   398: 'IGG_WARNING_WORD_01_BIT_5', class IGG Warnings, trigger "62_Warning_Data_IGG_WARNING_WORD_01" bit 13
   399: 'IGG_WARNING_WORD_01_BIT_6', class IGG Warnings, trigger "62_Warning_Data_IGG_WARNING_WORD_01" bit 14
   400: 'IGG_WARNING_WORD_01_BIT_7', class IGG Warnings, trigger "62_Warning_Data_IGG_WARNING_WORD_01" bit 15
   401: 'PIT-359 INLET CSW PRESSURE - LOW', class IGG Warnings, trigger "62_Warning_Data_IGG_WARNING_WORD_02" bit 0
   402: 'PIT-359 INLET CSW PRESSURE - HIGH', class IGG Warnings, trigger "62_Warning_Data_IGG_WARNING_WORD_02" bit 1
   403: 'PIT-316 OUTLET CSW PRESSURE - LOW', class IGG Warnings, trigger "62_Warning_Data_IGG_WARNING_WORD_02" bit 2
   404: 'PIT-316 OUTLET CSW PRESSURE - HIGH', class IGG Warnings, trigger "62_Warning_Data_IGG_WARNING_WORD_02" bit 3
   405: 'PIT-316 OUTLET CSW PRESSURE - LOW LOW', class IGG Warnings, trigger "62_Warning_Data_IGG_WARNING_WORD_02" bit 4
   406: 'PIT-316 OUTLET CSW PRESSURE - HIGH HIGH', class IGG Warnings, trigger "62_Warning_Data_IGG_WARNING_WORD_02" bit 5
   407: 'IGG_WARNING_WORD_02_BIT_14', class IGG Warnings, trigger "62_Warning_Data_IGG_WARNING_WORD_02" bit 6
   408: 'IGG_WARNING_WORD_02_BIT_15', class IGG Warnings, trigger "62_Warning_Data_IGG_WARNING_WORD_02" bit 7
   409: 'PIT-102 CA PRESSURE LOW', class IGG Warnings, trigger "62_Warning_Data_IGG_WARNING_WORD_02" bit 8
   410: 'PIT-102 CA PRESSURE HIGH', class IGG Warnings, trigger "62_Warning_Data_IGG_WARNING_WORD_02" bit 9
   411: 'TIT-401 IG TEMP HIGH', class IGG Warnings, trigger "62_Warning_Data_IGG_WARNING_WORD_02" bit 10
   412: 'PIT-402 IG OUTLET PRESSURE - LOW', class IGG Warnings, trigger "62_Warning_Data_IGG_WARNING_WORD_02" bit 11
   413: 'PIT-402 IG OUTLET PRESSURE - HIGH', class IGG Warnings, trigger "62_Warning_Data_IGG_WARNING_WORD_02" bit 12
   414: 'TIT-315 SHELL CSW TEMP - HIGH', class IGG Warnings, trigger "62_Warning_Data_IGG_WARNING_WORD_02" bit 13
   415: 'TIT-319 INLET CSW TEMP - HIGH', class IGG Warnings, trigger "62_Warning_Data_IGG_WARNING_WORD_02" bit 14
   416: 'TIT-360 OUTLET CSW TEMP - HIGH', class IGG Warnings, trigger "62_Warning_Data_IGG_WARNING_WORD_02" bit 15
   417: 'FD-001 FLAME - TRIPPED', class BC Warnings, trigger "62_Warning_Data_BC_WARNING_WORD_01" bit 0
   418: 'PIT-204 FUEL OIL INLET PRESSURE - LOW LOW', class BC Warnings, trigger "62_Warning_Data_BC_WARNING_WORD_01" bit 1
   419: 'PIT-204 FUEL OIL INLET PRESSURE - LOW', class BC Warnings, trigger "62_Warning_Data_BC_WARNING_WORD_01" bit 2
   420: 'PIT-204 FUEL OIL INLET PRESSURE - HIGH', class BC Warnings, trigger "62_Warning_Data_BC_WARNING_WORD_01" bit 3
   421: 'PIT-204 FUEL OIL INLET PRESSURE - HIGH HIGH', class BC Warnings, trigger "62_Warning_Data_BC_WARNING_WORD_01" bit 4
   422: 'PIT-204 FUEL OIL INLET PRESSURE - OUT OF RANGE', class BC Warnings, trigger "62_Warning_Data_BC_WARNING_WORD_01" bit 5
   423: 'BC_WARNING_WORD_01_BIT_14', class BC Warnings, trigger "62_Warning_Data_BC_WARNING_WORD_01" bit 6
   424: 'BC_WARNING_WORD_01_BIT_15', class BC Warnings, trigger "62_Warning_Data_BC_WARNING_WORD_01" bit 7
   425: 'BC_WARNING_WORD_01_BIT_0', class BC Warnings, trigger "62_Warning_Data_BC_WARNING_WORD_01" bit 8
   426: 'PIT-204 FUEL OIL INLET PRESSURE - LOW LOW', class BC Warnings, trigger "62_Warning_Data_BC_WARNING_WORD_01" bit 9
   427: 'PIT-204 FUEL OIL INLET PRESSURE - LOW', class BC Warnings, trigger "62_Warning_Data_BC_WARNING_WORD_01" bit 10
   428: 'PIT-204 FUEL OIL INLET PRESSURE - HIGH', class BC Warnings, trigger "62_Warning_Data_BC_WARNING_WORD_01" bit 11
   429: 'PIT-204 FUEL OIL INLET PRESSURE - HIGH HIGH', class BC Warnings, trigger "62_Warning_Data_BC_WARNING_WORD_01" bit 12
   430: 'PIT-204 FUEL OIL INLET PRESSURE - OUT OF RANGE', class BC Warnings, trigger "62_Warning_Data_BC_WARNING_WORD_01" bit 13
   431: 'FD-001 FLAME NOT DETECTED', class BC Warnings, trigger "62_Warning_Data_BC_WARNING_WORD_01" bit 14
   432: 'FD-001 FLAME NOT HEALTHY', class BC Warnings, trigger "62_Warning_Data_BC_WARNING_WORD_01" bit 15
   433: 'BC_WARNING_WORD_02_BIT_8', class BC Warnings, trigger "62_Warning_Data_BC_WARNING_WORD_02" bit 0
   434: 'TIT-202 FUEL OIL INLET TEMPERATURE - LOW LOW', class BC Warnings, trigger "62_Warning_Data_BC_WARNING_WORD_02" bit 1
   435: 'TIT-202 FUEL OIL INLET TEMPERATURE - LOW', class BC Warnings, trigger "62_Warning_Data_BC_WARNING_WORD_02" bit 2
   436: 'TIT-202 FUEL OIL INLET TEMPERATURE - HIGH', class BC Warnings, trigger "62_Warning_Data_BC_WARNING_WORD_02" bit 3
   437: 'TIT-202 FUEL OIL INLET TEMPERATURE - HIGH HIGH', class BC Warnings, trigger "62_Warning_Data_BC_WARNING_WORD_02" bit 4
   438: 'TIT-202 FUEL OIL INLET TEMPERATURE - OUT OF RANGE', class BC Warnings, trigger "62_Warning_Data_BC_WARNING_WORD_02" bit 5
   439: 'BC_WARNING_WORD_02_BIT_14', class BC Warnings, trigger "62_Warning_Data_BC_WARNING_WORD_02" bit 6
   440: 'BC_WARNING_WORD_02_BIT_15', class BC Warnings, trigger "62_Warning_Data_BC_WARNING_WORD_02" bit 7
   441: 'BC_WARNING_WORD_02_BIT_0', class BC Warnings, trigger "62_Warning_Data_BC_WARNING_WORD_02" bit 8
   442: 'TIT-202 IGG INLET FUEL TEMP - LOW LOW', class BC Warnings, trigger "62_Warning_Data_BC_WARNING_WORD_02" bit 9
   443: 'TIT-202 IGG INLET FUEL TEMP - LOW', class BC Warnings, trigger "62_Warning_Data_BC_WARNING_WORD_02" bit 10
   444: 'TIT-202 IGG INLET FUEL TEMP - HIGH', class BC Warnings, trigger "62_Warning_Data_BC_WARNING_WORD_02" bit 11
   445: 'TIT-202 IGG INLET FUEL TEMP - HIGH HIGH', class BC Warnings, trigger "62_Warning_Data_BC_WARNING_WORD_02" bit 12
   446: 'TIT-202 IGG INLET FUEL TEMP - OUT OF RANGE', class BC Warnings, trigger "62_Warning_Data_BC_WARNING_WORD_02" bit 13
   447: 'BC_WARNING_WORD_02_BIT_6', class BC Warnings, trigger "62_Warning_Data_BC_WARNING_WORD_02" bit 14
   448: 'BC_WARNING_WORD_02_BIT_7', class BC Warnings, trigger "62_Warning_Data_BC_WARNING_WORD_02" bit 15
   449: 'PIT-102 CA PRESSURE - LOW LOW', class IGG Warnings, trigger "62_Warning_Data_IGG_WARNING_WORD_03" bit 0
   450: 'PIT-102 CA PRESSURE - HIGH HIGH', class IGG Warnings, trigger "62_Warning_Data_IGG_WARNING_WORD_03" bit 1
   451: 'IGG WARNING', class IGG Warnings, trigger "62_Warning_Data_IGG_WARNING_WORD_03" bit 2
   452: 'PIT-402 IG OUTLET PRESSURE - LOW LOW', class IGG Warnings, trigger "62_Warning_Data_IGG_WARNING_WORD_03" bit 3
   453: 'PIT-402 IG OUTLET PRESSURE - HIGH HIGH', class IGG Warnings, trigger "62_Warning_Data_IGG_WARNING_WORD_03" bit 4
   454: 'TIT-315 SHELL CSW TEMP - HIGH HIGH', class IGG Warnings, trigger "62_Warning_Data_IGG_WARNING_WORD_03" bit 5
   455: 'TIT-319 INLET CSW TEMP - HIGH HIGH', class IGG Warnings, trigger "62_Warning_Data_IGG_WARNING_WORD_03" bit 6
   456: 'TIT-360 OUTLET CSW TEMP - HIGH HIGH', class IGG Warnings, trigger "62_Warning_Data_IGG_WARNING_WORD_03" bit 7
   457: 'PIT-112 IA PRESSURE- OUT OF RANGE', class IGG Warnings, trigger "62_Warning_Data_IGG_WARNING_WORD_03" bit 8
   458: 'PIT-113 FUEL PRESSURE TO MAIN BURNER - OUT OF RANGE', class IGG Warnings, trigger "62_Warning_Data_IGG_WARNING_WORD_03" bit 9
   459: 'PIT-102 CA PRESSURE - OUT OF RANGE', class IGG Warnings, trigger "62_Warning_Data_IGG_WARNING_WORD_03" bit 10
   460: 'TIT-401 IG TEMP - OUT OF RANGE', class IGG Warnings, trigger "62_Warning_Data_IGG_WARNING_WORD_03" bit 11
   461: 'PIT-402 IG VENT PRESSURE - OUT OF RANGE', class IGG Warnings, trigger "62_Warning_Data_IGG_WARNING_WORD_03" bit 12
   462: 'TIT-315 SHELL CSW TEMP - OUT OF RANGE', class IGG Warnings, trigger "62_Warning_Data_IGG_WARNING_WORD_03" bit 13
   463: 'TIT-319 INLET CSW TEMP - OUT OF RANGE', class IGG Warnings, trigger "62_Warning_Data_IGG_WARNING_WORD_03" bit 14
   464: 'TIT-360 OUTLET CSW TEMP - OUT OF RANGE', class IGG Warnings, trigger "62_Warning_Data_IGG_WARNING_WORD_03" bit 15
   465: 'INTERLOCKS NOT OK', class IGG Warnings, trigger "62_Warning_Data_IGG_WARNING_WORD_04" bit 0
   466: 'CHECK PIT-316 - WARNING', class IGG Warnings, trigger "62_Warning_Data_IGG_WARNING_WORD_04" bit 1
   467: 'CHECK PIT-102 - WARNING', class IGG Warnings, trigger "62_Warning_Data_IGG_WARNING_WORD_04" bit 2
   468: 'CHECK PIT-102 - WARNING II', class IGG Warnings, trigger "62_Warning_Data_IGG_WARNING_WORD_04" bit 3
   469: 'CHECK TIT-401 - WARNING', class IGG Warnings, trigger "62_Warning_Data_IGG_WARNING_WORD_04" bit 4
   470: 'CHECK TIT-319 - WARNING', class IGG Warnings, trigger "62_Warning_Data_IGG_WARNING_WORD_04" bit 5
   471: 'CHECK TIT-360 - WARNING', class IGG Warnings, trigger "62_Warning_Data_IGG_WARNING_WORD_04" bit 6
   472: 'E-500A TRIPPED', class IGG Warnings, trigger "62_Warning_Data_IGG_WARNING_WORD_04" bit 7
   473: 'E-500B TRIPPED', class IGG Warnings, trigger "62_Warning_Data_IGG_WARNING_WORD_04" bit 8
   474: 'PIT-359 INLET CSW PRESSURE - LOW LOW', class IGG Warnings, trigger "62_Warning_Data_IGG_WARNING_WORD_04" bit 9
   475: 'PIT-359 INLET CSW PRESSURE - HIGH HIGH', class IGG Warnings, trigger "62_Warning_Data_IGG_WARNING_WORD_04" bit 10
   476: 'PIT-359 INLET CSW PRESSURE - OUT OF RANGE', class IGG Warnings, trigger "62_Warning_Data_IGG_WARNING_WORD_04" bit 11
   477: 'PIT-316 OUTLET CSW PRESSURE - OUT OF RANGE', class IGG Warnings, trigger "62_Warning_Data_IGG_WARNING_WORD_04" bit 12
   478: 'PIT-112 IA PRESSURE - OUT OF RANGE', class IGG Warnings, trigger "62_Warning_Data_IGG_WARNING_WORD_04" bit 13
   479: 'IGG_WARNING_WORD_04_BIT_6', class IGG Warnings, trigger "62_Warning_Data_IGG_WARNING_WORD_04" bit 14
   480: 'IGG_WARNING_WORD_04_BIT_7', class IGG Warnings, trigger "62_Warning_Data_IGG_WARNING_WORD_04" bit 15
   481: 'BC_WARNING_WORD_03_BIT_8', class BC Warnings, trigger "62_Warning_Data_BC_WARNING_WORD_03" bit 0
   482: 'E-600 O2 ANALYSER CONTENT HIGH HIGH', class BC Warnings, trigger "62_Warning_Data_BC_WARNING_WORD_03" bit 1
   483: 'BC_WARNING_WORD_03_BIT_10', class BC Warnings, trigger "62_Warning_Data_BC_WARNING_WORD_03" bit 2
   484: 'BC_WARNING_WORD_03_BIT_11', class BC Warnings, trigger "62_Warning_Data_BC_WARNING_WORD_03" bit 3
   485: 'BC_WARNING_WORD_03_BIT_12', class BC Warnings, trigger "62_Warning_Data_BC_WARNING_WORD_03" bit 4
   486: 'BC_WARNING_WORD_03_BIT_13', class BC Warnings, trigger "62_Warning_Data_BC_WARNING_WORD_03" bit 5
   487: 'IGNITER POWER - NOT HEALTHY', class BC Warnings, trigger "62_Warning_Data_BC_WARNING_WORD_03" bit 6
   488: 'BC_WARNING_WORD_03_BIT_13', class BC Warnings, trigger "62_Warning_Data_BC_WARNING_WORD_03" bit 7
   489: 'BC_WARNING_WORD_03_BIT_0', class BC Warnings, trigger "62_Warning_Data_BC_WARNING_WORD_03" bit 8
   490: 'PIT-205 IGG MAIN FUEL PRESSURE - LOW', class BC Warnings, trigger "62_Warning_Data_BC_WARNING_WORD_03" bit 9
   491: 'PIT-205 IGG MAIN FUEL PRESSURE - LOW LOW', class BC Warnings, trigger "62_Warning_Data_BC_WARNING_WORD_03" bit 10
   492: 'PIT-205 IGG MAIN FUEL PRESSURE - HIGH', class BC Warnings, trigger "62_Warning_Data_BC_WARNING_WORD_03" bit 11
   493: 'PIT-205 IGG MAIN FUEL PRESSURE - HIGH HIGH', class BC Warnings, trigger "62_Warning_Data_BC_WARNING_WORD_03" bit 12
   494: 'PIT-205 IGG MAIN FUEL PRESSURE - OUT OF RANGE', class BC Warnings, trigger "62_Warning_Data_BC_WARNING_WORD_03" bit 13
   495: 'E-131 IA COMPRESSOR - WARNING', class BC Warnings, trigger "62_Warning_Data_BC_WARNING_WORD_03" bit 14
   496: 'E-131 IA COMPRESSOR - NOT RUNNING', class BC Warnings, trigger "62_Warning_Data_BC_WARNING_WORD_03" bit 15
   497: 'CHECK PIT-112 IA PRESSURE - WARNING', class BC Warnings, trigger "62_Warning_Data_BC_WARNING_WORD_04" bit 0
   498: 'CHECK PIT-204 FUEL OIL INLET PRESSURE - WARNING', class BC Warnings, trigger "62_Warning_Data_BC_WARNING_WORD_04" bit 1
   499: 'CHECK FS-123 PILOT AIR FLOW - WARNING', class BC Warnings, trigger "62_Warning_Data_BC_WARNING_WORD_04" bit 2
   500: 'CHECK FS-115 MAIN BURNER ATOMISING AIR FLOW - WARNING', class BC Warnings, trigger "62_Warning_Data_BC_WARNING_WORD_04" bit 3
   501: 'CHECK FS-317 IGG JACKET COOLING WATER FLOW - WARNING', class BC Warnings, trigger "62_Warning_Data_BC_WARNING_WORD_04" bit 4
   502: 'SOOT SYSTEM POWER - NOT HEALTHY', class BC Warnings, trigger "62_Warning_Data_BC_WARNING_WORD_04" bit 5
   503: 'SOOT SYSTEM OPACITY - HIGH', class BC Warnings, trigger "62_Warning_Data_BC_WARNING_WORD_04" bit 6
   504: 'SOOT SYSTEM - OUT OF RANGE', class BC Warnings, trigger "62_Warning_Data_BC_WARNING_WORD_04" bit 7
   505: 'BC_INTERLOCKS NOT OK', class BC Warnings, trigger "62_Warning_Data_BC_WARNING_WORD_04" bit 8
   506: 'PIT-112 INLET IA PRESSURE - LOW LOW', class BC Warnings, trigger "62_Warning_Data_BC_WARNING_WORD_04" bit 9
   507: 'PIT-112 INLET IA PRESSURE - LOW', class BC Warnings, trigger "62_Warning_Data_BC_WARNING_WORD_04" bit 10
   508: 'PIT-112 INLET IA PRESSURE - HIGH', class BC Warnings, trigger "62_Warning_Data_BC_WARNING_WORD_04" bit 11
   509: 'PIT-112 INLET IA PRESSURE - HIGH HIGH', class BC Warnings, trigger "62_Warning_Data_BC_WARNING_WORD_04" bit 12
   510: 'PIT-112 INLET IA PRESSURE - OUT OF RANGE', class BC Warnings, trigger "62_Warning_Data_BC_WARNING_WORD_04" bit 13
   511: 'CHECK FS-317 IGG JACKET COOLING WATER FLOW - WARNING', class BC Warnings, trigger "62_Warning_Data_BC_WARNING_WORD_04" bit 14
   512: 'CHECK FS-320 REAR MATRIX COOLING WATER FLOW - WARNING', class BC Warnings, trigger "62_Warning_Data_BC_WARNING_WORD_04" bit 15
   513: 'IGG HMI LOST COMUNICATION', class IGG Warnings, trigger "62_Warning_Data_IGG_WARNING_WORD_05" bit 0
   514: 'CCR HMI LOST COMUNICATION', class IGG Warnings, trigger "62_Warning_Data_IGG_WARNING_WORD_05" bit 1
   515: 'BRIGE HMI LOST COMUNICATION', class IGG Warnings, trigger "62_Warning_Data_IGG_WARNING_WORD_05" bit 2
   516: 'PIT-402 CA PRESSURE - LOW LOW', class IGG Warnings, trigger "62_Warning_Data_IGG_WARNING_WORD_05" bit 3
   517: 'PIT-402 CA PRESSURE - HIGH HIGH', class IGG Warnings, trigger "62_Warning_Data_IGG_WARNING_WORD_05" bit 4
   518: 'TIT-315 SHELL CSW TEMP - HIGH HIGH', class IGG Warnings, trigger "62_Warning_Data_IGG_WARNING_WORD_05" bit 5
   519: 'TIT-319 INLET CSW TEMP - HIGH HIGH', class IGG Warnings, trigger "62_Warning_Data_IGG_WARNING_WORD_05" bit 6
   520: 'TIT-360 OUTLET CSW TEMP - HIGH HIGH', class IGG Warnings, trigger "62_Warning_Data_IGG_WARNING_WORD_05" bit 7
   521: 'BC PLC POWER NOT HEALTHY', class IGG Warnings, trigger "62_Warning_Data_IGG_WARNING_WORD_05" bit 8
   522: 'CONTROLS POWER SUPPLY - NOT HEALTHY', class IGG Warnings, trigger "62_Warning_Data_IGG_WARNING_WORD_05" bit 9
   523: 'IGG POWER SUPPLY - NOT HEALTHY', class IGG Warnings, trigger "62_Warning_Data_IGG_WARNING_WORD_05" bit 10
   524: 'BC POWER SUPPLY - NOT HEALTHY', class IGG Warnings, trigger "62_Warning_Data_IGG_WARNING_WORD_05" bit 11
   525: 'BACKUP 24VDC POWER SUPPLY - NOT HEALTHY', class IGG Warnings, trigger "62_Warning_Data_IGG_WARNING_WORD_05" bit 12
   526: 'IGG VENTILATION POWER - NOT HEALTHY', class IGG Warnings, trigger "62_Warning_Data_IGG_WARNING_WORD_05" bit 13
   527: 'MCCP VENTILATION POWER - NOT HEALTHY', class IGG Warnings, trigger "62_Warning_Data_IGG_WARNING_WORD_05" bit 14
   528: 'TIT-360 OUTLET CSW TEMP - HIGH HIGH', class IGG Warnings, trigger "62_Warning_Data_IGG_WARNING_WORD_05" bit 15
   529: 'PIT-359 INLET CSW PRESSURE - LOW LOW', class IGG Warnings, trigger "62_Warning_Data_IGG_WARNING_WORD_06" bit 0
   530: 'PIT-359 INLET CSW PRESSURE - HIGH HIGH', class IGG Warnings, trigger "62_Warning_Data_IGG_WARNING_WORD_06" bit 1
   531: 'IGG_WARNING_WORD_06_BIT_10', class IGG Warnings, trigger "62_Warning_Data_IGG_WARNING_WORD_06" bit 2
   532: 'IGG_WARNING_WORD_06_BIT_11', class IGG Warnings, trigger "62_Warning_Data_IGG_WARNING_WORD_06" bit 3
   533: 'IGG_WARNING_WORD_06_BIT_12', class IGG Warnings, trigger "62_Warning_Data_IGG_WARNING_WORD_06" bit 4
   534: 'IGG_WARNING_WORD_06_BIT_13', class IGG Warnings, trigger "62_Warning_Data_IGG_WARNING_WORD_06" bit 5
   535: 'IGG_WARNING_WORD_06_BIT_14', class IGG Warnings, trigger "62_Warning_Data_IGG_WARNING_WORD_06" bit 6
   536: 'IGG_WARNING_WORD_06_BIT_15', class IGG Warnings, trigger "62_Warning_Data_IGG_WARNING_WORD_06" bit 7
   537: 'IGG_WARNING_WORD_06_BIT_0', class IGG Warnings, trigger "62_Warning_Data_IGG_WARNING_WORD_06" bit 8
   538: 'IGG_WARNING_WORD_06_BIT_1', class IGG Warnings, trigger "62_Warning_Data_IGG_WARNING_WORD_06" bit 9
   539: 'IGG_WARNING_WORD_06_BIT_2', class IGG Warnings, trigger "62_Warning_Data_IGG_WARNING_WORD_06" bit 10
   540: 'IGG_WARNING_WORD_06_BIT_3', class IGG Warnings, trigger "62_Warning_Data_IGG_WARNING_WORD_06" bit 11
   541: 'IGG_WARNING_WORD_06_BIT_4', class IGG Warnings, trigger "62_Warning_Data_IGG_WARNING_WORD_06" bit 12
   542: 'IGG_WARNING_WORD_06_BIT_5', class IGG Warnings, trigger "62_Warning_Data_IGG_WARNING_WORD_06" bit 13
   543: 'IGG_WARNING_WORD_06_BIT_6', class IGG Warnings, trigger "62_Warning_Data_IGG_WARNING_WORD_06" bit 14
   544: 'IGG_WARNING_WORD_06_BIT_7', class IGG Warnings, trigger "62_Warning_Data_IGG_WARNING_WORD_06" bit 15
   545: 'BC_WARNING_WORD_05_BIT_8', class BC Warnings, trigger "62_Warning_Data_BC_WARNING_WORD_05" bit 0
   546: 'BC_WARNING_WORD_05_BIT_9', class BC Warnings, trigger "62_Warning_Data_BC_WARNING_WORD_05" bit 1
   547: 'BC_WARNING_WORD_05_BIT_10', class BC Warnings, trigger "62_Warning_Data_BC_WARNING_WORD_05" bit 2
   548: 'BC_WARNING_WORD_05_BIT_11', class BC Warnings, trigger "62_Warning_Data_BC_WARNING_WORD_05" bit 3
   549: 'BC_WARNING_WORD_05_BIT_12', class BC Warnings, trigger "62_Warning_Data_BC_WARNING_WORD_05" bit 4
   550: 'BC_WARNING_WORD_05_BIT_13', class BC Warnings, trigger "62_Warning_Data_BC_WARNING_WORD_05" bit 5
   551: 'BC_WARNING_WORD_05_BIT_14', class BC Warnings, trigger "62_Warning_Data_BC_WARNING_WORD_05" bit 6
   552: 'BC_WARNING_WORD_05_BIT_15', class BC Warnings, trigger "62_Warning_Data_BC_WARNING_WORD_05" bit 7
   553: 'BC_WARNING_WORD_05_BIT_0', class BC Warnings, trigger "62_Warning_Data_BC_WARNING_WORD_05" bit 8
   554: 'PIT-113 IGG MAIN ATOM AIR PRESSURE - LOW LOW', class BC Warnings, trigger "62_Warning_Data_BC_WARNING_WORD_05" bit 9
   555: 'PIT-113 IGG MAIN ATOM AIR PRESSURE - LOW', class BC Warnings, trigger "62_Warning_Data_BC_WARNING_WORD_05" bit 10
   556: 'PIT-113 IGG MAIN ATOM AIR PRESSURE - HIGH', class BC Warnings, trigger "62_Warning_Data_BC_WARNING_WORD_05" bit 11
   557: 'PIT-113 IGG MAIN ATOM AIR PRESSURE - HIGH HIGH', class BC Warnings, trigger "62_Warning_Data_BC_WARNING_WORD_05" bit 12
   558: 'PIT-113 IGG MAIN ATOM AIR PRESSURE - OUT OF RANGE', class BC Warnings, trigger "62_Warning_Data_BC_WARNING_WORD_05" bit 13
   559: 'BC_WARNING_WORD', class BC Warnings, trigger "62_Warning_Data_BC_WARNING_WORD_05" bit 14
   560: 'BC_WARNING WORD', class BC Warnings, trigger "62_Warning_Data_BC_WARNING_WORD_05" bit 15
   561: 'INTERLOCKS NOT OK', class BC Warnings, trigger "62_Warning_Data_BC_WARNING_WORD_06" bit 0
   562: 'BC_WARNING_WORD_06_BIT_9', class BC Warnings, trigger "62_Warning_Data_BC_WARNING_WORD_06" bit 1
   563: 'BC_WARNING_WORD_06_BIT_10', class BC Warnings, trigger "62_Warning_Data_BC_WARNING_WORD_06" bit 2
   564: 'BC_WARNING_WORD_06_BIT_11', class BC Warnings, trigger "62_Warning_Data_BC_WARNING_WORD_06" bit 3
   565: 'BC_WARNING_WORD_06_BIT_12', class BC Warnings, trigger "62_Warning_Data_BC_WARNING_WORD_06" bit 4
   566: 'BC_WARNING_WORD_06_BIT_13', class BC Warnings, trigger "62_Warning_Data_BC_WARNING_WORD_06" bit 5
   567: 'BC_WARNING_WORD_06_BIT_14', class BC Warnings, trigger "62_Warning_Data_BC_WARNING_WORD_06" bit 6
   568: 'BC_WARNING_WORD_06_BIT_15', class BC Warnings, trigger "62_Warning_Data_BC_WARNING_WORD_06" bit 7
   569: 'INTERLOCKS NOT OK', class BC Warnings, trigger "62_Warning_Data_BC_WARNING_WORD_06" bit 8
   570: 'BC_WARNING_WORD_06_BIT_1', class BC Warnings, trigger "62_Warning_Data_BC_WARNING_WORD_06" bit 9
   571: 'BC_WARNING_WORD_06_BIT_2', class BC Warnings, trigger "62_Warning_Data_BC_WARNING_WORD_06" bit 10
   572: 'BC_WARNING_WORD_06_BIT_3', class BC Warnings, trigger "62_Warning_Data_BC_WARNING_WORD_06" bit 11
   573: 'BC_WARNING_WORD_06_BIT_4', class BC Warnings, trigger "62_Warning_Data_BC_WARNING_WORD_06" bit 12
   574: 'BC_WARNING_WORD_06_BIT_5', class BC Warnings, trigger "62_Warning_Data_BC_WARNING_WORD_06" bit 13
   575: 'BC_WARNING_WORD_06_BIT_6', class BC Warnings, trigger "62_Warning_Data_BC_WARNING_WORD_06" bit 14
   576: 'BC_WARNING_WORD_06_BIT_7', class BC Warnings, trigger "62_Warning_Data_BC_WARNING_WORD_06" bit 15
   577: 'BC_WARNING_WORD_05_BIT_8', class BC Warnings bit 0
   1000: 'E-400 - FAULT', class GCU Alarms, trigger "60_Alarm_Data_GCU_ALARM_WORD_01" bit 0
   1001: 'GCU_ALARM_WORD_01_BIT_9', class GCU Alarms, trigger "60_Alarm_Data_GCU_ALARM_WORD_01" bit 1
   1002: 'GCU_ALARM_WORD_01_BIT_10', class GCU Alarms, trigger "60_Alarm_Data_GCU_ALARM_WORD_01" bit 2
   1003: 'GCU_ALARM_WORD_01_BIT_11', class GCU Alarms, trigger "60_Alarm_Data_GCU_ALARM_WORD_01" bit 3
   1004: 'GCU_ALARM_WORD_01_BIT_12', class GCU Alarms, trigger "60_Alarm_Data_GCU_ALARM_WORD_01" bit 4
   1005: 'GCU_ALARM_WORD_01_BIT_13', class GCU Alarms, trigger "60_Alarm_Data_GCU_ALARM_WORD_01" bit 5
   1006: 'GCU_ALARM_WORD_01_BIT_14', class GCU Alarms, trigger "60_Alarm_Data_GCU_ALARM_WORD_01" bit 6
   1007: 'GCU_ALARM_WORD_01_BIT_15', class GCU Alarms, trigger "60_Alarm_Data_GCU_ALARM_WORD_01" bit 7
   1008: 'BWT PANEL E-STOP PRESSED', class GCU Alarms, trigger "60_Alarm_Data_GCU_ALARM_WORD_01" bit 8
   1009: 'GCU SLAVE PLC HEART BEAT MISSING', class GCU Alarms, trigger "60_Alarm_Data_GCU_ALARM_WORD_01" bit 9
   1010: 'GCU BWTS AUTO INTERLOCKS NOT OK', class GCU Alarms, trigger "60_Alarm_Data_GCU_ALARM_WORD_01" bit 10
   1011: 'LIT-304 GCU TANK LEVEL HIGH HIGH', class GCU Alarms, trigger "60_Alarm_Data_GCU_ALARM_WORD_01" bit 11
   1012: 'LIT-304 LIQUID LEVEL LOW LOW', class GCU Alarms, trigger "60_Alarm_Data_GCU_ALARM_WORD_01" bit 12
   1013: 'P-303 FRESH RECIRCULATION PUMP - TRIPPED', class GCU Alarms, trigger "60_Alarm_Data_GCU_ALARM_WORD_01" bit 13
   1014: 'P-304 FRESH WATER BOOSTER PUMP - TRIPPED', class GCU Alarms, trigger "60_Alarm_Data_GCU_ALARM_WORD_01" bit 14
   1015: 'E-400 PROCESS GAS COMPRESSOR - TRIPPED', class GCU Alarms, trigger "60_Alarm_Data_GCU_ALARM_WORD_01" bit 15
   1016: 'PIT-353 RECIRCULATION FRESH WATER PRESSURE HIGH HIGH', class GCU Alarms, trigger "60_Alarm_Data_GCU_ALARM_WORD_02" bit 0
   1017: 'PIT-416 GAS TO DECK PRESSURE LOW LOW', class GCU Alarms, trigger "60_Alarm_Data_GCU_ALARM_WORD_02" bit 1
   1018: 'PIT-416 GAS TO DECK PRESSURE HIGH HIGH', class GCU Alarms, trigger "60_Alarm_Data_GCU_ALARM_WORD_02" bit 2
   1019: 'PIT-358 FRESH WATER INLET PRESSURE - LOW LOW', class GCU Alarms, trigger "60_Alarm_Data_GCU_ALARM_WORD_02" bit 3
   1020: 'PIT-358 FRESH WATER INLET PRESSURE - HIGH HIGH', class GCU Alarms, trigger "60_Alarm_Data_GCU_ALARM_WORD_02" bit 4
   1021: 'PIT-348 COOLING SEA WATER TO E-300 PRESSURE - LOW LOW', class GCU Alarms, trigger "60_Alarm_Data_GCU_ALARM_WORD_02" bit 5
   1022: 'PIT-348 COOLING SEA WATER TO E-300 PRESSURE HIGH HIGH', class GCU Alarms, trigger "60_Alarm_Data_GCU_ALARM_WORD_02" bit 6
   1023: 'GCU_ALARM_WORD_02_BIT_15', class GCU Alarms, trigger "60_Alarm_Data_GCU_ALARM_WORD_02" bit 7
   1024: 'FS-332 COOLING SEA WATER TO E-300 - LOW FLOW', class GCU Alarms, trigger "60_Alarm_Data_GCU_ALARM_WORD_02" bit 8
   1025: 'PIT-348 COOLING SEA WATER TO E-300 PRESSURE - LOW LOW', class GCU Alarms, trigger "60_Alarm_Data_GCU_ALARM_WORD_02" bit 9
   1026: 'PIT-348 COOLING SEA WATER TO E-300 PRESSURE - HIGH HIGH', class GCU Alarms, trigger "60_Alarm_Data_GCU_ALARM_WORD_02" bit 10
   1027: 'FS-350 FRESH WATER COOLING TO GCU FLOW - LOW FLOW', class GCU Alarms, trigger "60_Alarm_Data_GCU_ALARM_WORD_02" bit 11
   1028: 'GCU_ALARM_WORD_02_BIT_4', class GCU Alarms, trigger "60_Alarm_Data_GCU_ALARM_WORD_02" bit 12
   1029: 'TIT-002 - HIGH HIGH', class GCU Alarms, trigger "60_Alarm_Data_GCU_ALARM_WORD_02" bit 13
   1030: 'PIT-002 - HIGH HIGH', class GCU Alarms, trigger "60_Alarm_Data_GCU_ALARM_WORD_02" bit 14
   1031: 'PIT-353 RECIRCULATION FRESH WATER PRESSURE - LOW LOW', class GCU Alarms, trigger "60_Alarm_Data_GCU_ALARM_WORD_02" bit 15
   1032: 'PIT-353 RECIRCULATION FRESH WATER PRESSURE - HIGH HIGH', class GCU Alarms, trigger "60_Alarm_Data_GCU_ALARM_WORD_03" bit 0
   1033: 'PIT-416 GAS TO DECK PRESSURE - LOW LOW', class GCU Alarms, trigger "60_Alarm_Data_GCU_ALARM_WORD_03" bit 1
   1034: 'PIT-416 GAS TO DECK PRESSURE - HIGH HIGH', class GCU Alarms, trigger "60_Alarm_Data_GCU_ALARM_WORD_03" bit 2
   1035: 'PIT-358 FRESH WATER INLET PRESSURE - LOW LOW', class GCU Alarms, trigger "60_Alarm_Data_GCU_ALARM_WORD_03" bit 3
   1036: 'PIT-358 FRESH WATER INLET PRESSURE - HIGH HIGH', class GCU Alarms, trigger "60_Alarm_Data_GCU_ALARM_WORD_03" bit 4
   1037: 'PIT-348 COOLING SEA WATER TO E-300 PRESSURE - LOW LOW', class GCU Alarms, trigger "60_Alarm_Data_GCU_ALARM_WORD_03" bit 5
   1038: 'PIT-348 COOLING SEA WATER TO E-300 PRESSURE - HIGH HIGH', class GCU Alarms, trigger "60_Alarm_Data_GCU_ALARM_WORD_03" bit 6
   1039: 'GCU_ALARM_WORD_03_BIT_15', class GCU Alarms, trigger "60_Alarm_Data_GCU_ALARM_WORD_03" bit 7
   1040: 'GCU_ALARM_WORD_03_BIT_0', class GCU Alarms, trigger "60_Alarm_Data_GCU_ALARM_WORD_03" bit 8
   1041: 'GCU_ALARM_WORD_03_BIT_1', class GCU Alarms, trigger "60_Alarm_Data_GCU_ALARM_WORD_03" bit 9
   1042: 'GCU_ALARM_WORD_03_BIT_2', class GCU Alarms, trigger "60_Alarm_Data_GCU_ALARM_WORD_03" bit 10
   1043: 'GCU_ALARM_WORD_03_BIT_3', class GCU Alarms, trigger "60_Alarm_Data_GCU_ALARM_WORD_03" bit 11
   1044: 'GCU_ALARM_WORD_03_BIT_4', class GCU Alarms, trigger "60_Alarm_Data_GCU_ALARM_WORD_03" bit 12
   1045: 'GCU_ALARM_WORD_03_BIT_5', class GCU Alarms, trigger "60_Alarm_Data_GCU_ALARM_WORD_03" bit 13
   1046: 'GCU_ALARM_WORD_03_BIT_6', class GCU Alarms, trigger "60_Alarm_Data_GCU_ALARM_WORD_03" bit 14
   1047: 'GCU_ALARM_WORD_03_BIT_7', class GCU Alarms, trigger "60_Alarm_Data_GCU_ALARM_WORD_03" bit 15
   1048: 'GCU_ALARM_WORD_04_BIT_8', class GCU Alarms, trigger "60_Alarm_Data_GCU_ALARM_WORD_04" bit 0
   1049: 'GCU_ALARM_WORD_04_BIT_9', class GCU Alarms, trigger "60_Alarm_Data_GCU_ALARM_WORD_04" bit 1
   1050: 'GCU_ALARM_WORD_04_BIT_10', class GCU Alarms, trigger "60_Alarm_Data_GCU_ALARM_WORD_04" bit 2
   1051: 'GCU_ALARM_WORD_04_BIT_11', class GCU Alarms, trigger "60_Alarm_Data_GCU_ALARM_WORD_04" bit 3
   1052: 'GCU_ALARM_WORD_04_BIT_12', class GCU Alarms, trigger "60_Alarm_Data_GCU_ALARM_WORD_04" bit 4
   1053: 'GCU_ALARM_WORD_04_BIT_13', class GCU Alarms, trigger "60_Alarm_Data_GCU_ALARM_WORD_04" bit 5
   1054: 'GCU_ALARM_WORD_04_BIT_14', class GCU Alarms, trigger "60_Alarm_Data_GCU_ALARM_WORD_04" bit 6
   1055: 'GCU_ALARM_WORD_04_BIT_15', class GCU Alarms, trigger "60_Alarm_Data_GCU_ALARM_WORD_04" bit 7
   1056: 'CV-341 GCU DRAIN VALVE - FAULT', class GCU Alarms, trigger "60_Alarm_Data_GCU_ALARM_WORD_04" bit 8
   1057: 'CV-358 FRESH WATER SUPPLY LINE CONTROL VALVE - FAULT', class GCU Alarms, trigger "60_Alarm_Data_GCU_ALARM_WORD_04" bit 9
   1058: 'CV-406 DECK ISOLATION VALVE - FAULT', class GCU Alarms, trigger "60_Alarm_Data_GCU_ALARM_WORD_04" bit 10
   1059: 'CV-407 DECK MAIN ISOLATION VALVE 1 - FAULT', class GCU Alarms, trigger "60_Alarm_Data_GCU_ALARM_WORD_04" bit 11
   1060: 'CV-409 DOUBLE BLOCK AND BLEED VENT VALVE - FAULT', class GCU Alarms, trigger "60_Alarm_Data_GCU_ALARM_WORD_04" bit 12
   1061: 'CV-411 DECK MAIN ISOLATION VALVE 2 - FAULT', class GCU Alarms, trigger "60_Alarm_Data_GCU_ALARM_WORD_04" bit 13
   1062: 'CV-441 PGC AIR INLET VALVE - FAULT', class GCU Alarms, trigger "60_Alarm_Data_GCU_ALARM_WORD_04" bit 14
   1063: 'GCU_ALARM_WORD_04_BIT_7', class GCU Alarms, trigger "60_Alarm_Data_GCU_ALARM_WORD_04" bit 15
   1064: 'GCU_ALARM_WORD_05_BIT_8', class GCU Alarms, trigger "60_Alarm_Data_GCU_ALARM_WORD_05" bit 0
   1065: 'GCU_ALARM_WORD_05_BIT_9', class GCU Alarms, trigger "60_Alarm_Data_GCU_ALARM_WORD_05" bit 1
   1066: 'GCU_ALARM_WORD_05_BIT_10', class GCU Alarms, trigger "60_Alarm_Data_GCU_ALARM_WORD_05" bit 2
   1067: 'GCU_ALARM_WORD_05_BIT_11', class GCU Alarms, trigger "60_Alarm_Data_GCU_ALARM_WORD_05" bit 3
   1068: 'GCU_ALARM_WORD_05_BIT_12', class GCU Alarms, trigger "60_Alarm_Data_GCU_ALARM_WORD_05" bit 4
   1069: 'GCU_ALARM_WORD_05_BIT_13', class GCU Alarms, trigger "60_Alarm_Data_GCU_ALARM_WORD_05" bit 5
   1070: 'GCU_ALARM_WORD_05_BIT_14', class GCU Alarms, trigger "60_Alarm_Data_GCU_ALARM_WORD_05" bit 6
   1071: 'GCU_ALARM_WORD_05_BIT_15', class GCU Alarms, trigger "60_Alarm_Data_GCU_ALARM_WORD_05" bit 7
   1072: 'GCU_ALARM_WORD_05_BIT_0', class GCU Alarms, trigger "60_Alarm_Data_GCU_ALARM_WORD_05" bit 8
   1073: 'GCU_ALARM_WORD_05_BIT_1', class GCU Alarms, trigger "60_Alarm_Data_GCU_ALARM_WORD_05" bit 9
   1074: 'GCU_ALARM_WORD_05_BIT_2', class GCU Alarms, trigger "60_Alarm_Data_GCU_ALARM_WORD_05" bit 10
   1075: 'GCU_ALARM_WORD_05_BIT_3', class GCU Alarms, trigger "60_Alarm_Data_GCU_ALARM_WORD_05" bit 11
   1076: 'GCU_ALARM_WORD_05_BIT_4', class GCU Alarms, trigger "60_Alarm_Data_GCU_ALARM_WORD_05" bit 12
   1077: 'GCU_ALARM_WORD_05_BIT_5', class GCU Alarms, trigger "60_Alarm_Data_GCU_ALARM_WORD_05" bit 13
   1078: 'GCU_ALARM_WORD_05_BIT_6', class GCU Alarms, trigger "60_Alarm_Data_GCU_ALARM_WORD_05" bit 14
   1079: 'GCU_ALARM_WORD_05_BIT_7', class GCU Alarms, trigger "60_Alarm_Data_GCU_ALARM_WORD_05" bit 15
   1080: 'GCU_ALARM_WORD_06_BIT_8', class GCU Alarms, trigger "60_Alarm_Data_GCU_ALARM_WORD_06" bit 0
   1081: 'GCU_ALARM_WORD_06_BIT_9', class GCU Alarms, trigger "60_Alarm_Data_GCU_ALARM_WORD_06" bit 1
   1082: 'GCU_ALARM_WORD_06_BIT_10', class GCU Alarms, trigger "60_Alarm_Data_GCU_ALARM_WORD_06" bit 2
   1083: 'GCU_ALARM_WORD_06_BIT_11', class GCU Alarms, trigger "60_Alarm_Data_GCU_ALARM_WORD_06" bit 3
   1084: 'GCU_ALARM_WORD_06_BIT_12', class GCU Alarms, trigger "60_Alarm_Data_GCU_ALARM_WORD_06" bit 4
   1085: 'GCU_ALARM_WORD_06_BIT_13', class GCU Alarms, trigger "60_Alarm_Data_GCU_ALARM_WORD_06" bit 5
   1086: 'GCU_ALARM_WORD_06_BIT_14', class GCU Alarms, trigger "60_Alarm_Data_GCU_ALARM_WORD_06" bit 6
   1087: 'GCU_ALARM_WORD_06_BIT_15', class GCU Alarms, trigger "60_Alarm_Data_GCU_ALARM_WORD_06" bit 7
   1088: 'GCU_ALARM_WORD_06_BIT_0', class GCU Alarms, trigger "60_Alarm_Data_GCU_ALARM_WORD_06" bit 8
   1089: 'GCU_ALARM_WORD_06_BIT_1', class GCU Alarms, trigger "60_Alarm_Data_GCU_ALARM_WORD_06" bit 9
   1090: 'GCU_ALARM_WORD_06_BIT_2', class GCU Alarms, trigger "60_Alarm_Data_GCU_ALARM_WORD_06" bit 10
   1091: 'GCU_ALARM_WORD_06_BIT_3', class GCU Alarms, trigger "60_Alarm_Data_GCU_ALARM_WORD_06" bit 11
   1092: 'GCU_ALARM_WORD_06_BIT_4', class GCU Alarms, trigger "60_Alarm_Data_GCU_ALARM_WORD_06" bit 12
   1093: 'GCU_ALARM_WORD_06_BIT_5', class GCU Alarms, trigger "60_Alarm_Data_GCU_ALARM_WORD_06" bit 13
   1094: 'GCU_ALARM_WORD_06_BIT_6', class GCU Alarms, trigger "60_Alarm_Data_GCU_ALARM_WORD_06" bit 14
   1095: 'GCU_ALARM_WORD_06_BIT_7', class GCU Alarms, trigger "60_Alarm_Data_GCU_ALARM_WORD_06" bit 15
   1096: 'GCU_ALARM_WORD_07_BIT_8', class GCU Alarms, trigger "60_Alarm_Data_GCU_ALARM_WORD_07" bit 0
   1097: 'GCU_ALARM_WORD_07_BIT_9', class GCU Alarms, trigger "60_Alarm_Data_GCU_ALARM_WORD_07" bit 1
   1098: 'GCU_ALARM_WORD_07_BIT_10', class GCU Alarms, trigger "60_Alarm_Data_GCU_ALARM_WORD_07" bit 2
   1099: 'GCU_ALARM_WORD_07_BIT_11', class GCU Alarms, trigger "60_Alarm_Data_GCU_ALARM_WORD_07" bit 3
   1100: 'GCU_ALARM_WORD_07_BIT_12', class GCU Alarms, trigger "60_Alarm_Data_GCU_ALARM_WORD_07" bit 4
   1101: 'GCU_ALARM_WORD_07_BIT_13', class GCU Alarms, trigger "60_Alarm_Data_GCU_ALARM_WORD_07" bit 5
   1102: 'GCU_ALARM_WORD_07_BIT_14', class GCU Alarms, trigger "60_Alarm_Data_GCU_ALARM_WORD_07" bit 6
   1103: 'GCU_ALARM_WORD_07_BIT_15', class GCU Alarms, trigger "60_Alarm_Data_GCU_ALARM_WORD_07" bit 7
   1104: 'GCU_ALARM_WORD_07_BIT_0', class GCU Alarms, trigger "60_Alarm_Data_GCU_ALARM_WORD_07" bit 8
   1105: 'GCU_ALARM_WORD_07_BIT_1', class GCU Alarms, trigger "60_Alarm_Data_GCU_ALARM_WORD_07" bit 9
   1106: 'GCU_ALARM_WORD_07_BIT_2', class GCU Alarms, trigger "60_Alarm_Data_GCU_ALARM_WORD_07" bit 10
   1107: 'GCU_ALARM_WORD_07_BIT_3', class GCU Alarms, trigger "60_Alarm_Data_GCU_ALARM_WORD_07" bit 11
   1108: 'GCU_ALARM_WORD_07_BIT_4', class GCU Alarms, trigger "60_Alarm_Data_GCU_ALARM_WORD_07" bit 12
   1109: 'GCU_ALARM_WORD_07_BIT_5', class GCU Alarms, trigger "60_Alarm_Data_GCU_ALARM_WORD_07" bit 13
   1110: 'GCU_ALARM_WORD_07_BIT_6', class GCU Alarms, trigger "60_Alarm_Data_GCU_ALARM_WORD_07" bit 14
   1111: 'GCU_ALARM_WORD_07_BIT_7', class GCU Alarms, trigger "60_Alarm_Data_GCU_ALARM_WORD_07" bit 15
   1112: 'GCU_ALARM_WORD_08_BIT_8', class GCU Alarms, trigger "60_Alarm_Data_GCU_ALARM_WORD_08" bit 0
   1113: 'GCU_ALARM_WORD_08_BIT_9', class GCU Alarms, trigger "60_Alarm_Data_GCU_ALARM_WORD_08" bit 1
   1114: 'GCU_ALARM_WORD_08_BIT_10', class GCU Alarms, trigger "60_Alarm_Data_GCU_ALARM_WORD_08" bit 2
   1115: 'GCU_ALARM_WORD_08_BIT_11', class GCU Alarms, trigger "60_Alarm_Data_GCU_ALARM_WORD_08" bit 3
   1116: 'GCU_ALARM_WORD_08_BIT_12', class GCU Alarms, trigger "60_Alarm_Data_GCU_ALARM_WORD_08" bit 4
   1117: 'GCU_ALARM_WORD_08_BIT_13', class GCU Alarms, trigger "60_Alarm_Data_GCU_ALARM_WORD_08" bit 5
